      { S7_Templates := "SrcType := Int" } LE_Contact(in1 := "100_GCU_AUTO_SEQ_DB".CRNT_STEP, in2 := 470)
   END_RUNG wire#w1
   // the same network as SCL:
   "Setpoint Override_DB"(Enable := ("100_GCU_AUTO_SEQ_DB".CRNT_STEP >= 290) AND ("100_GCU_AUTO_SEQ_DB".CRNT_STEP <= 470),   // "Setpoint Override"
                          "Activate Temp Prot" := "80_From_HMI"."TT002 Target Protection",
                          Temperature := "12_AI_Data".E_400_TE002_SCALED,
                          "Temperature Setpoint" := "84_Setpoints".E400_TT002_HighHigh,
                          "Temperature Tolerance" := "84_Setpoints"."E-400 TT002 Tolerance",
                          "Activate Press Prot" := "80_From_HMI"."PT002 Target Protection",
                          Pressure := "12_AI_Data".E_400_PT002_SCALED,
                          "Pressure Setpoint" := "84_Setpoints".E400_PT002_High,
                          "Pressure Tolerance" := "84_Setpoints"."E-400 PT002 Tolerance",
                          "Pressure Target" := "84_Setpoints".PIT416_Target,
                          "Pressure Safe Target" := "84_Setpoints".PIT416_Target_Safe,
                          "Activate Tank Change Prot" := "80_From_HMI"."Tank Close Protection",
                          "Tank Change TimeOut" := "84_Setpoints"."Tank Close TimeOut",
                          "Pressure Safe Override" => "84_Setpoints".PIT416_Target_Safe,
                          ENO => #_w1);
   IF #_w1 AND "Setpoint Override_DB"."Set Pressure" THEN
       "19_AUTO_CMNDS_Data".PIT416_CMND_Target := "Setpoint Override_DB"."Pressure Target Override";
   END_IF;
END_REGION

REGION Network 6: PIT416 Target Ramp
   RUNG wire#powerrail
      { S7_Templates := "[SrcType := Real, DestType := DInt]" } Convert(in := "86_Times".PIT416_TRGT_RMP_TIME, out => "68_Sys_Status_Data"."PIT416_TRGT_RMP_TIME D_INT")
      Mul(in1 := "68_Sys_Status_Data"."PIT416_TRGT_RMP_TIME D_INT", in2 := 1000, out => "RAMP_DB"."Time span")
      "RAMP_DB"(Start := wire#w1, "Time span" :=, "Minimum Value" := "12_AI_Data".PIT_416_SCALED, "Maximum Value" := "84_Setpoints".PIT416_Target, Value =>, "Ramp Done" =>)
      I_Contact( "Setpoint Override_DB"."Set Pressure" )
      Move(in := "RAMP_DB".Value, out1 => "19_AUTO_CMNDS_Data".PIT416_CMND_Target)
   END_RUNG
   RUNG wire#powerrail
      { S7_Templates := "SrcType := Int" } GE_Contact(in1 := "100_GCU_AUTO_SEQ_DB".CRNT_STEP, in2 := 290)
      { S7_Templates := "SrcType := Int" } LT_Contact(in1 := "100_GCU_AUTO_SEQ_DB".CRNT_STEP, in2 := 450)
   END_RUNG wire#w1
   // the same network as SCL:
   "68_Sys_Status_Data"."PIT416_TRGT_RMP_TIME D_INT" := REAL_TO_DINT("86_Times".PIT416_TRGT_RMP_TIME);
   "RAMP_DB"."Time span" := "68_Sys_Status_Data"."PIT416_TRGT_RMP_TIME D_INT" * 1000;
   "RAMP_DB"(Start := ("100_GCU_AUTO_SEQ_DB".CRNT_STEP >= 290) AND ("100_GCU_AUTO_SEQ_DB".CRNT_STEP < 450),   // "RAMP"
             "Minimum Value" := "12_AI_Data".PIT_416_SCALED,
             "Maximum Value" := "84_Setpoints".PIT416_Target,
             ENO => #_w1);
   IF #_w1 AND NOT "Setpoint Override_DB"."Set Pressure" THEN
       "19_AUTO_CMNDS_Data".PIT416_CMND_Target := "RAMP_DB".Value;
   END_IF;
END_REGION
END_FUNCTION

FUNCTION "150_GCU_LCL_CNTRL" : Void   // FC150, LAD
TITLE = GCU Local Control
{ S7_Optimized_Access := 'TRUE' }
AUTHOR : JRS
VERSION : 0.1
// For automatic control of the GCU from the HMI and not the BWTS or BTCS
   VAR_TEMP   // added for the SCL form of the ladder/FBD networks
      _w1 : Bool;
   END_VAR
BEGIN

REGION Network 1: System Ok For Local Control
   // Valves at initial etc
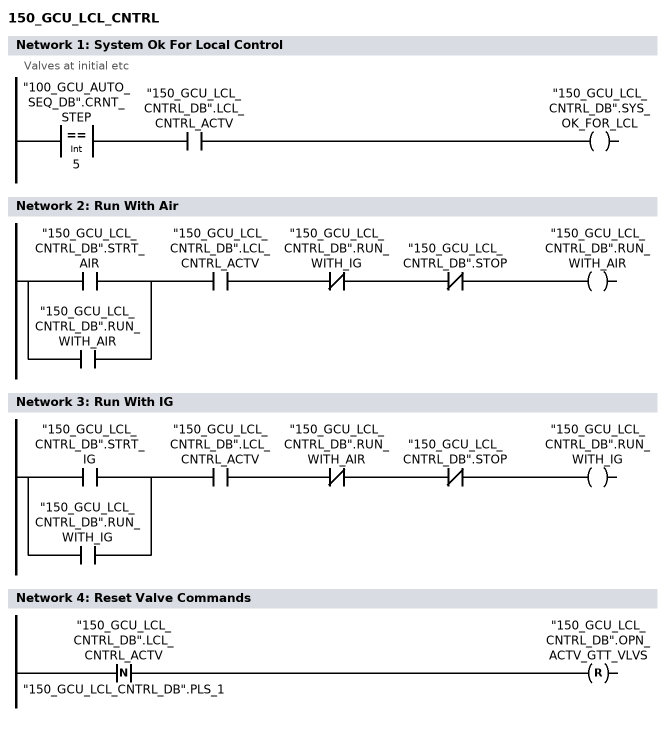
   RUNG wire#powerrail
      { S7_Templates := "SrcType := Int" } EQ_Contact(in1 := "100_GCU_AUTO_SEQ_DB".CRNT_STEP, in2 := 5)
      Contact( "150_GCU_LCL_CNTRL_DB".LCL_CNTRL_ACTV )
      Coil( "150_GCU_LCL_CNTRL_DB".SYS_OK_FOR_LCL )
   END_RUNG
   // the same network as SCL:
   "150_GCU_LCL_CNTRL_DB".SYS_OK_FOR_LCL := ("100_GCU_AUTO_SEQ_DB".CRNT_STEP = 5) AND "150_GCU_LCL_CNTRL_DB".LCL_CNTRL_ACTV;
END_REGION

REGION Network 2: Run With Air
   RUNG wire#powerrail
      Contact( "150_GCU_LCL_CNTRL_DB".STRT_AIR )
      wire#w1
      Contact( "150_GCU_LCL_CNTRL_DB".LCL_CNTRL_ACTV )
      I_Contact( "150_GCU_LCL_CNTRL_DB".RUN_WITH_IG )
      I_Contact( "150_GCU_LCL_CNTRL_DB".STOP )
      Coil( "150_GCU_LCL_CNTRL_DB".RUN_WITH_AIR )
   END_RUNG
   RUNG wire#powerrail
      Contact( "150_GCU_LCL_CNTRL_DB".RUN_WITH_AIR )
   END_RUNG wire#w1
   // the same network as SCL:
   "150_GCU_LCL_CNTRL_DB".RUN_WITH_AIR := ("150_GCU_LCL_CNTRL_DB".STRT_AIR OR "150_GCU_LCL_CNTRL_DB".RUN_WITH_AIR) AND "150_GCU_LCL_CNTRL_DB".LCL_CNTRL_ACTV AND NOT "150_GCU_LCL_CNTRL_DB".RUN_WITH_IG AND NOT "150_GCU_LCL_CNTRL_DB".STOP;
END_REGION

REGION Network 3: Run With IG
   RUNG wire#powerrail
      Contact( "150_GCU_LCL_CNTRL_DB".STRT_IG )
      wire#w1
      Contact( "150_GCU_LCL_CNTRL_DB".LCL_CNTRL_ACTV )
      I_Contact( "150_GCU_LCL_CNTRL_DB".RUN_WITH_AIR )
      I_Contact( "150_GCU_LCL_CNTRL_DB".STOP )
      Coil( "150_GCU_LCL_CNTRL_DB".RUN_WITH_IG )
   END_RUNG
   RUNG wire#powerrail
      Contact( "150_GCU_LCL_CNTRL_DB".RUN_WITH_IG )
   END_RUNG wire#w1
   // the same network as SCL:
   "150_GCU_LCL_CNTRL_DB".RUN_WITH_IG := ("150_GCU_LCL_CNTRL_DB".STRT_IG OR "150_GCU_LCL_CNTRL_DB".RUN_WITH_IG) AND "150_GCU_LCL_CNTRL_DB".LCL_CNTRL_ACTV AND NOT "150_GCU_LCL_CNTRL_DB".RUN_WITH_AIR AND NOT "150_GCU_LCL_CNTRL_DB".STOP;
END_REGION

REGION Network 4: Reset Valve Commands
   RUNG wire#powerrail
      N_Contact(operand := "150_GCU_LCL_CNTRL_DB".LCL_CNTRL_ACTV, bit := "150_GCU_LCL_CNTRL_DB".PLS_1)
      R_Coil( "150_GCU_LCL_CNTRL_DB".OPN_ACTV_GTT_VLVS )
   END_RUNG
   // the same network as SCL:
   #_w1 := NOT "150_GCU_LCL_CNTRL_DB".LCL_CNTRL_ACTV AND "150_GCU_LCL_CNTRL_DB".PLS_1;   // falling edge of "150_GCU_LCL_CNTRL_DB".LCL_CNTRL_ACTV
   "150_GCU_LCL_CNTRL_DB".PLS_1 := "150_GCU_LCL_CNTRL_DB".LCL_CNTRL_ACTV;
   IF #_w1 THEN "150_GCU_LCL_CNTRL_DB".OPN_ACTV_GTT_VLVS := FALSE; END_IF;
END_REGION
END_FUNCTION

// folder: 1000 - 1999 BWT System Control/1060 - 1089 Alarm & Valve Status Handling

FUNCTION "1060_ALARMS_TO_WORDS" : Void   // FC1060, LAD
TITLE = Alarm Processing
{ S7_Optimized_Access := 'TRUE' }
AUTHOR : JRS
VERSION : 0.1
// To determine alarm conditions
BEGIN

REGION Network 1: DB64 DBX18.0 = TX425/426 Tank 1 pH Low Alarm
   // BWTS_ALARM_WORD_10_BIT_0
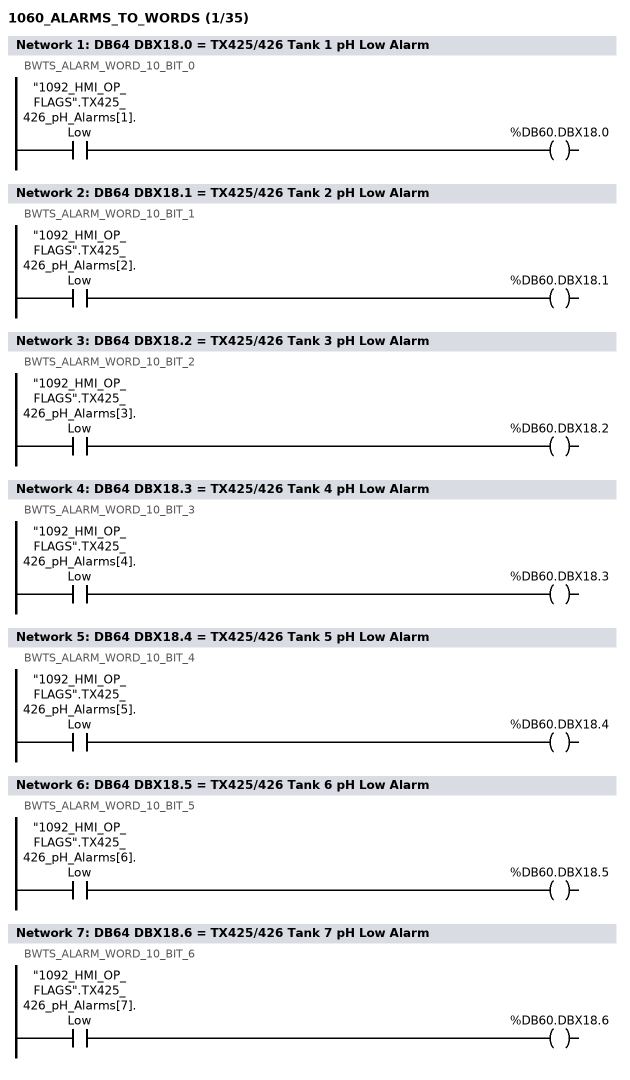
   RUNG wire#powerrail
      Contact( "1092_HMI_OP_FLAGS".TX425_426_pH_Alarms[1].Low )
      Coil( %DB60.DBX18.0 )
   END_RUNG
   // the same network as SCL:
   %DB60.DBX18.0 := "1092_HMI_OP_FLAGS".TX425_426_pH_Alarms[1].Low;
END_REGION

REGION Network 2: DB64 DBX18.1 = TX425/426 Tank 2 pH Low Alarm
   // BWTS_ALARM_WORD_10_BIT_1
   RUNG wire#powerrail
      Contact( "1092_HMI_OP_FLAGS".TX425_426_pH_Alarms[2].Low )
      Coil( %DB60.DBX18.1 )
   END_RUNG
   // the same network as SCL:
   %DB60.DBX18.1 := "1092_HMI_OP_FLAGS".TX425_426_pH_Alarms[2].Low;
END_REGION

REGION Network 3: DB64 DBX18.2 = TX425/426 Tank 3 pH Low Alarm
   // BWTS_ALARM_WORD_10_BIT_2
   RUNG wire#powerrail
      Contact( "1092_HMI_OP_FLAGS".TX425_426_pH_Alarms[3].Low )
      Coil( %DB60.DBX18.2 )
   END_RUNG
   // the same network as SCL:
   %DB60.DBX18.2 := "1092_HMI_OP_FLAGS".TX425_426_pH_Alarms[3].Low;
END_REGION

REGION Network 4: DB64 DBX18.3 = TX425/426 Tank 4 pH Low Alarm
   // BWTS_ALARM_WORD_10_BIT_3
   RUNG wire#powerrail
      Contact( "1092_HMI_OP_FLAGS".TX425_426_pH_Alarms[4].Low )
      Coil( %DB60.DBX18.3 )
   END_RUNG
   // the same network as SCL:
   %DB60.DBX18.3 := "1092_HMI_OP_FLAGS".TX425_426_pH_Alarms[4].Low;
END_REGION

REGION Network 5: DB64 DBX18.4 = TX425/426 Tank 5 pH Low Alarm
   // BWTS_ALARM_WORD_10_BIT_4
   RUNG wire#powerrail
      Contact( "1092_HMI_OP_FLAGS".TX425_426_pH_Alarms[5].Low )
      Coil( %DB60.DBX18.4 )
   END_RUNG
   // the same network as SCL:
   %DB60.DBX18.4 := "1092_HMI_OP_FLAGS".TX425_426_pH_Alarms[5].Low;
END_REGION

REGION Network 6: DB64 DBX18.5 = TX425/426 Tank 6 pH Low Alarm
   // BWTS_ALARM_WORD_10_BIT_5
   RUNG wire#powerrail
      Contact( "1092_HMI_OP_FLAGS".TX425_426_pH_Alarms[6].Low )
      Coil( %DB60.DBX18.5 )
   END_RUNG
   // the same network as SCL:
   %DB60.DBX18.5 := "1092_HMI_OP_FLAGS".TX425_426_pH_Alarms[6].Low;
END_REGION

REGION Network 7: DB64 DBX18.6 = TX425/426 Tank 7 pH Low Alarm
   // BWTS_ALARM_WORD_10_BIT_6
   RUNG wire#powerrail
      Contact( "1092_HMI_OP_FLAGS".TX425_426_pH_Alarms[7].Low )
      Coil( %DB60.DBX18.6 )
   END_RUNG
   // the same network as SCL:
   %DB60.DBX18.6 := "1092_HMI_OP_FLAGS".TX425_426_pH_Alarms[7].Low;
END_REGION

REGION Network 8: DB64 DBX18.7 = TX425/426 Tank 8 pH Low Alarm
   // BWTS_ALARM_WORD_10_BIT_7
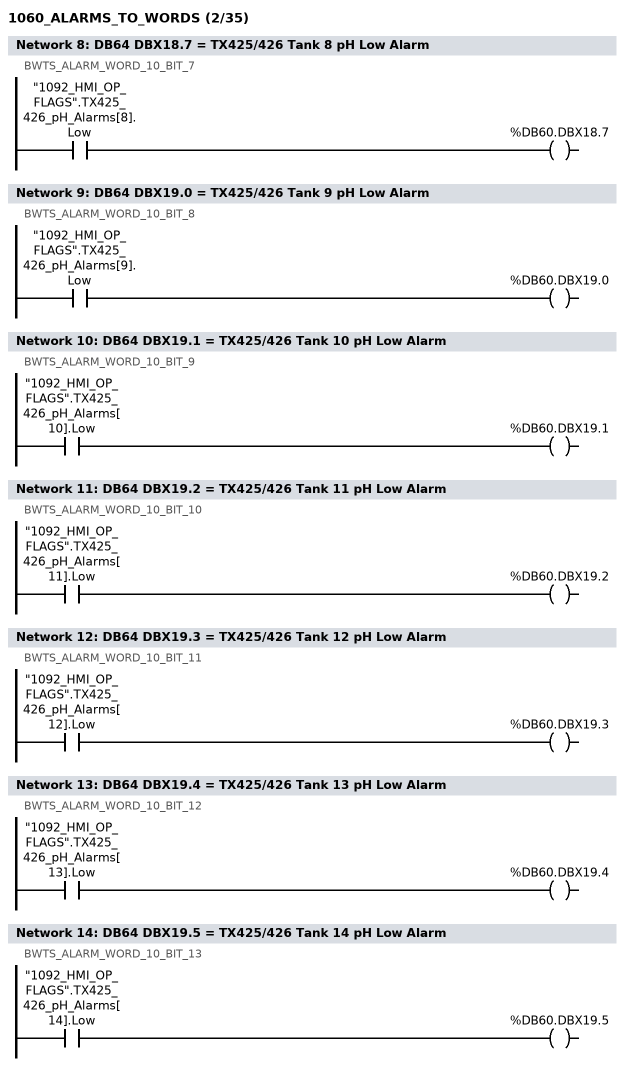
   RUNG wire#powerrail
      Contact( "1092_HMI_OP_FLAGS".TX425_426_pH_Alarms[8].Low )
      Coil( %DB60.DBX18.7 )
   END_RUNG
   // the same network as SCL:
   %DB60.DBX18.7 := "1092_HMI_OP_FLAGS".TX425_426_pH_Alarms[8].Low;
END_REGION

REGION Network 9: DB64 DBX19.0 = TX425/426 Tank 9 pH Low Alarm
   // BWTS_ALARM_WORD_10_BIT_8
   RUNG wire#powerrail
      Contact( "1092_HMI_OP_FLAGS".TX425_426_pH_Alarms[9].Low )
      Coil( %DB60.DBX19.0 )
   END_RUNG
   // the same network as SCL:
   %DB60.DBX19.0 := "1092_HMI_OP_FLAGS".TX425_426_pH_Alarms[9].Low;
END_REGION

REGION Network 10: DB64 DBX19.1 = TX425/426 Tank 10 pH Low Alarm
   // BWTS_ALARM_WORD_10_BIT_9
   RUNG wire#powerrail
      Contact( "1092_HMI_OP_FLAGS".TX425_426_pH_Alarms[10].Low )
      Coil( %DB60.DBX19.1 )
   END_RUNG
   // the same network as SCL:
   %DB60.DBX19.1 := "1092_HMI_OP_FLAGS".TX425_426_pH_Alarms[10].Low;
END_REGION

REGION Network 11: DB64 DBX19.2 = TX425/426 Tank 11 pH Low Alarm
   // BWTS_ALARM_WORD_10_BIT_10
   RUNG wire#powerrail
      Contact( "1092_HMI_OP_FLAGS".TX425_426_pH_Alarms[11].Low )
      Coil( %DB60.DBX19.2 )
   END_RUNG
   // the same network as SCL:
   %DB60.DBX19.2 := "1092_HMI_OP_FLAGS".TX425_426_pH_Alarms[11].Low;
END_REGION

REGION Network 12: DB64 DBX19.3 = TX425/426 Tank 12 pH Low Alarm
   // BWTS_ALARM_WORD_10_BIT_11
   RUNG wire#powerrail
      Contact( "1092_HMI_OP_FLAGS".TX425_426_pH_Alarms[12].Low )
      Coil( %DB60.DBX19.3 )
   END_RUNG
   // the same network as SCL:
   %DB60.DBX19.3 := "1092_HMI_OP_FLAGS".TX425_426_pH_Alarms[12].Low;
END_REGION

REGION Network 13: DB64 DBX19.4 = TX425/426 Tank 13 pH Low Alarm
   // BWTS_ALARM_WORD_10_BIT_12
   RUNG wire#powerrail
      Contact( "1092_HMI_OP_FLAGS".TX425_426_pH_Alarms[13].Low )
      Coil( %DB60.DBX19.4 )
   END_RUNG
   // the same network as SCL:
   %DB60.DBX19.4 := "1092_HMI_OP_FLAGS".TX425_426_pH_Alarms[13].Low;
END_REGION

REGION Network 14: DB64 DBX19.5 = TX425/426 Tank 14 pH Low Alarm
   // BWTS_ALARM_WORD_10_BIT_13
   RUNG wire#powerrail
      Contact( "1092_HMI_OP_FLAGS".TX425_426_pH_Alarms[14].Low )
      Coil( %DB60.DBX19.5 )
   END_RUNG
   // the same network as SCL:
   %DB60.DBX19.5 := "1092_HMI_OP_FLAGS".TX425_426_pH_Alarms[14].Low;
END_REGION

REGION Network 16: DB64 DBX20.0 = TX427/428 Tank 1 DO Low Alarm
   // BWTS_ALARM_WORD_11_BIT_0
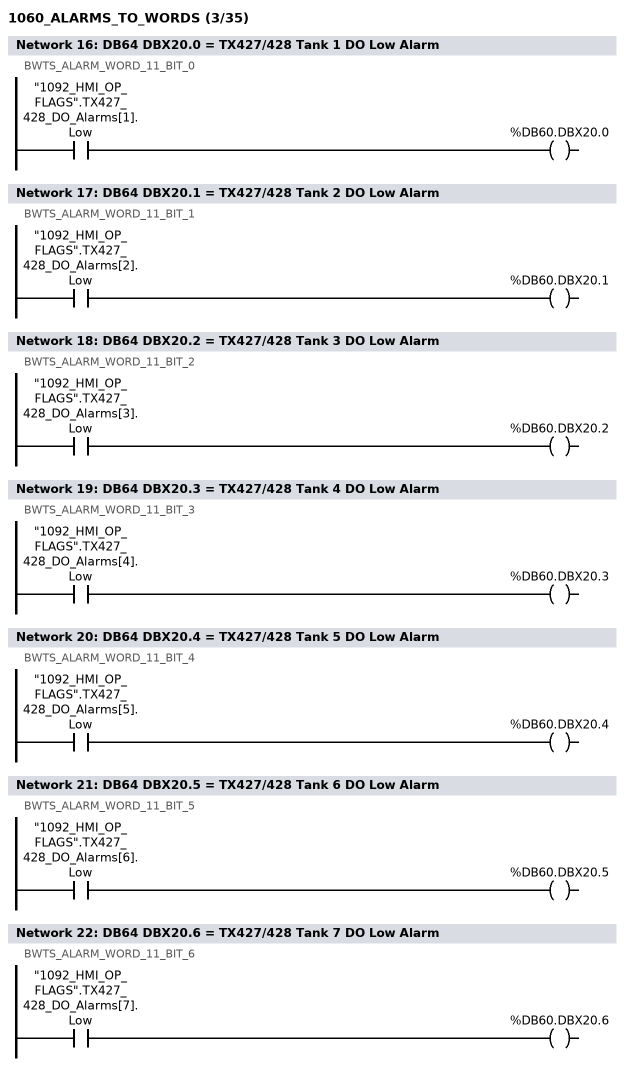
   RUNG wire#powerrail
      Contact( "1092_HMI_OP_FLAGS".TX427_428_DO_Alarms[1].Low )
      Coil( %DB60.DBX20.0 )
   END_RUNG
   // the same network as SCL:
   %DB60.DBX20.0 := "1092_HMI_OP_FLAGS".TX427_428_DO_Alarms[1].Low;
END_REGION

REGION Network 17: DB64 DBX20.1 = TX427/428 Tank 2 DO Low Alarm
   // BWTS_ALARM_WORD_11_BIT_1
   RUNG wire#powerrail
      Contact( "1092_HMI_OP_FLAGS".TX427_428_DO_Alarms[2].Low )
      Coil( %DB60.DBX20.1 )
   END_RUNG
   // the same network as SCL:
   %DB60.DBX20.1 := "1092_HMI_OP_FLAGS".TX427_428_DO_Alarms[2].Low;
END_REGION

REGION Network 18: DB64 DBX20.2 = TX427/428 Tank 3 DO Low Alarm
   // BWTS_ALARM_WORD_11_BIT_2
   RUNG wire#powerrail
      Contact( "1092_HMI_OP_FLAGS".TX427_428_DO_Alarms[3].Low )
      Coil( %DB60.DBX20.2 )
   END_RUNG
   // the same network as SCL:
   %DB60.DBX20.2 := "1092_HMI_OP_FLAGS".TX427_428_DO_Alarms[3].Low;
END_REGION

REGION Network 19: DB64 DBX20.3 = TX427/428 Tank 4 DO Low Alarm
   // BWTS_ALARM_WORD_11_BIT_3
   RUNG wire#powerrail
      Contact( "1092_HMI_OP_FLAGS".TX427_428_DO_Alarms[4].Low )
      Coil( %DB60.DBX20.3 )
   END_RUNG
   // the same network as SCL:
   %DB60.DBX20.3 := "1092_HMI_OP_FLAGS".TX427_428_DO_Alarms[4].Low;
END_REGION

REGION Network 20: DB64 DBX20.4 = TX427/428 Tank 5 DO Low Alarm
   // BWTS_ALARM_WORD_11_BIT_4
   RUNG wire#powerrail
      Contact( "1092_HMI_OP_FLAGS".TX427_428_DO_Alarms[5].Low )
      Coil( %DB60.DBX20.4 )
   END_RUNG
   // the same network as SCL:
   %DB60.DBX20.4 := "1092_HMI_OP_FLAGS".TX427_428_DO_Alarms[5].Low;
END_REGION

REGION Network 21: DB64 DBX20.5 = TX427/428 Tank 6 DO Low Alarm
   // BWTS_ALARM_WORD_11_BIT_5
   RUNG wire#powerrail
      Contact( "1092_HMI_OP_FLAGS".TX427_428_DO_Alarms[6].Low )
      Coil( %DB60.DBX20.5 )
   END_RUNG
   // the same network as SCL:
   %DB60.DBX20.5 := "1092_HMI_OP_FLAGS".TX427_428_DO_Alarms[6].Low;
END_REGION

REGION Network 22: DB64 DBX20.6 = TX427/428 Tank 7 DO Low Alarm
   // BWTS_ALARM_WORD_11_BIT_6
   RUNG wire#powerrail
      Contact( "1092_HMI_OP_FLAGS".TX427_428_DO_Alarms[7].Low )
      Coil( %DB60.DBX20.6 )
   END_RUNG
   // the same network as SCL:
   %DB60.DBX20.6 := "1092_HMI_OP_FLAGS".TX427_428_DO_Alarms[7].Low;
END_REGION

REGION Network 23: DB64 DBX20.7 = TX427/428 Tank 8 DO Low Alarm
   // BWTS_ALARM_WORD_11_BIT_7
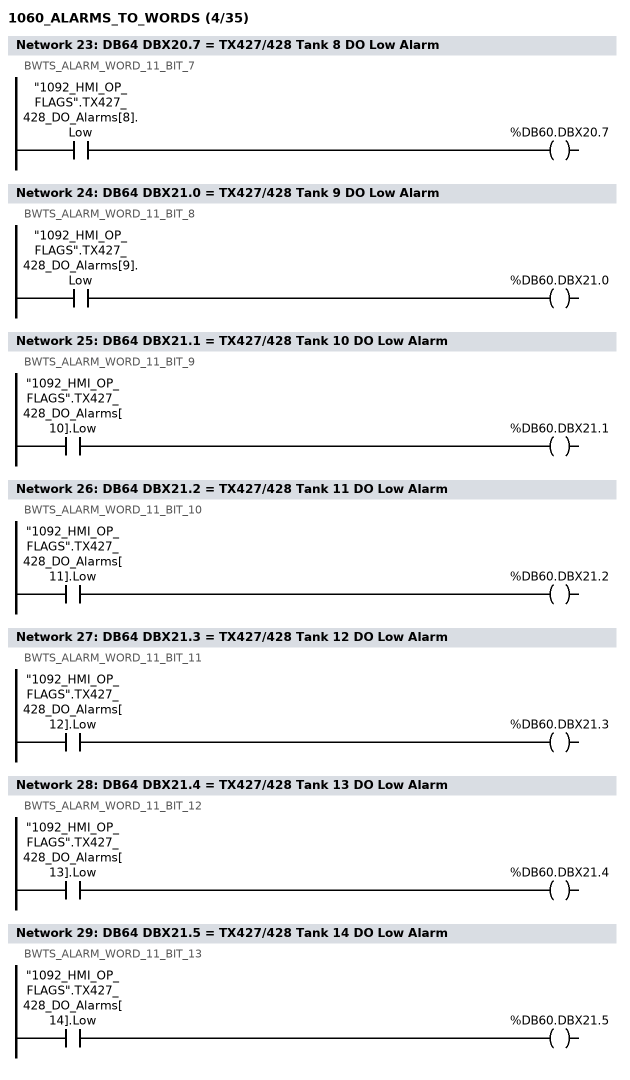
   RUNG wire#powerrail
      Contact( "1092_HMI_OP_FLAGS".TX427_428_DO_Alarms[8].Low )
      Coil( %DB60.DBX20.7 )
   END_RUNG
   // the same network as SCL:
   %DB60.DBX20.7 := "1092_HMI_OP_FLAGS".TX427_428_DO_Alarms[8].Low;
END_REGION

REGION Network 24: DB64 DBX21.0 = TX427/428 Tank 9 DO Low Alarm
   // BWTS_ALARM_WORD_11_BIT_8
   RUNG wire#powerrail
      Contact( "1092_HMI_OP_FLAGS".TX427_428_DO_Alarms[9].Low )
      Coil( %DB60.DBX21.0 )
   END_RUNG
   // the same network as SCL:
   %DB60.DBX21.0 := "1092_HMI_OP_FLAGS".TX427_428_DO_Alarms[9].Low;
END_REGION

REGION Network 25: DB64 DBX21.1 = TX427/428 Tank 10 DO Low Alarm
   // BWTS_ALARM_WORD_11_BIT_9
   RUNG wire#powerrail
      Contact( "1092_HMI_OP_FLAGS".TX427_428_DO_Alarms[10].Low )
      Coil( %DB60.DBX21.1 )
   END_RUNG
   // the same network as SCL:
   %DB60.DBX21.1 := "1092_HMI_OP_FLAGS".TX427_428_DO_Alarms[10].Low;
END_REGION

REGION Network 26: DB64 DBX21.2 = TX427/428 Tank 11 DO Low Alarm
   // BWTS_ALARM_WORD_11_BIT_10
   RUNG wire#powerrail
      Contact( "1092_HMI_OP_FLAGS".TX427_428_DO_Alarms[11].Low )
      Coil( %DB60.DBX21.2 )
   END_RUNG
   // the same network as SCL:
   %DB60.DBX21.2 := "1092_HMI_OP_FLAGS".TX427_428_DO_Alarms[11].Low;
END_REGION

REGION Network 27: DB64 DBX21.3 = TX427/428 Tank 12 DO Low Alarm
   // BWTS_ALARM_WORD_11_BIT_11
   RUNG wire#powerrail
      Contact( "1092_HMI_OP_FLAGS".TX427_428_DO_Alarms[12].Low )
      Coil( %DB60.DBX21.3 )
   END_RUNG
   // the same network as SCL:
   %DB60.DBX21.3 := "1092_HMI_OP_FLAGS".TX427_428_DO_Alarms[12].Low;
END_REGION

REGION Network 28: DB64 DBX21.4 = TX427/428 Tank 13 DO Low Alarm
   // BWTS_ALARM_WORD_11_BIT_12
   RUNG wire#powerrail
      Contact( "1092_HMI_OP_FLAGS".TX427_428_DO_Alarms[13].Low )
      Coil( %DB60.DBX21.4 )
   END_RUNG
   // the same network as SCL:
   %DB60.DBX21.4 := "1092_HMI_OP_FLAGS".TX427_428_DO_Alarms[13].Low;
END_REGION

REGION Network 29: DB64 DBX21.5 = TX427/428 Tank 14 DO Low Alarm
   // BWTS_ALARM_WORD_11_BIT_13
   RUNG wire#powerrail
      Contact( "1092_HMI_OP_FLAGS".TX427_428_DO_Alarms[14].Low )
      Coil( %DB60.DBX21.5 )
   END_RUNG
   // the same network as SCL:
   %DB60.DBX21.5 := "1092_HMI_OP_FLAGS".TX427_428_DO_Alarms[14].Low;
END_REGION

REGION Network 31: DB64 DBX22.0 = USD Flow Tank 1 Low Low
   // BWTS_ALARM_WORD_12_BIT_0
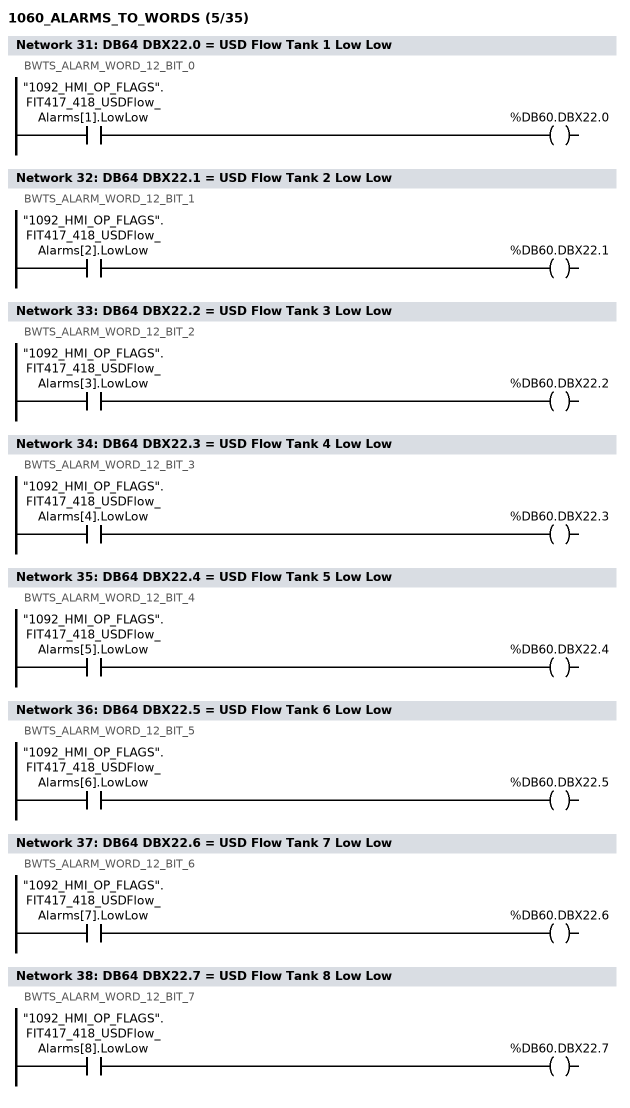
   RUNG wire#powerrail
      Contact( "1092_HMI_OP_FLAGS".FIT417_418_USDFlow_Alarms[1].LowLow )
      Coil( %DB60.DBX22.0 )
   END_RUNG
   // the same network as SCL:
   %DB60.DBX22.0 := "1092_HMI_OP_FLAGS".FIT417_418_USDFlow_Alarms[1].LowLow;
END_REGION

REGION Network 32: DB64 DBX22.1 = USD Flow Tank 2 Low Low
   // BWTS_ALARM_WORD_12_BIT_1
   RUNG wire#powerrail
      Contact( "1092_HMI_OP_FLAGS".FIT417_418_USDFlow_Alarms[2].LowLow )
      Coil( %DB60.DBX22.1 )
   END_RUNG
   // the same network as SCL:
   %DB60.DBX22.1 := "1092_HMI_OP_FLAGS".FIT417_418_USDFlow_Alarms[2].LowLow;
END_REGION

REGION Network 33: DB64 DBX22.2 = USD Flow Tank 3 Low Low
   // BWTS_ALARM_WORD_12_BIT_2
   RUNG wire#powerrail
      Contact( "1092_HMI_OP_FLAGS".FIT417_418_USDFlow_Alarms[3].LowLow )
      Coil( %DB60.DBX22.2 )
   END_RUNG
   // the same network as SCL:
   %DB60.DBX22.2 := "1092_HMI_OP_FLAGS".FIT417_418_USDFlow_Alarms[3].LowLow;
END_REGION

REGION Network 34: DB64 DBX22.3 = USD Flow Tank 4 Low Low
   // BWTS_ALARM_WORD_12_BIT_3
   RUNG wire#powerrail
      Contact( "1092_HMI_OP_FLAGS".FIT417_418_USDFlow_Alarms[4].LowLow )
      Coil( %DB60.DBX22.3 )
   END_RUNG
   // the same network as SCL:
   %DB60.DBX22.3 := "1092_HMI_OP_FLAGS".FIT417_418_USDFlow_Alarms[4].LowLow;
END_REGION

REGION Network 35: DB64 DBX22.4 = USD Flow Tank 5 Low Low
   // BWTS_ALARM_WORD_12_BIT_4
   RUNG wire#powerrail
      Contact( "1092_HMI_OP_FLAGS".FIT417_418_USDFlow_Alarms[5].LowLow )
      Coil( %DB60.DBX22.4 )
   END_RUNG
   // the same network as SCL:
   %DB60.DBX22.4 := "1092_HMI_OP_FLAGS".FIT417_418_USDFlow_Alarms[5].LowLow;
END_REGION

REGION Network 36: DB64 DBX22.5 = USD Flow Tank 6 Low Low
   // BWTS_ALARM_WORD_12_BIT_5
   RUNG wire#powerrail
      Contact( "1092_HMI_OP_FLAGS".FIT417_418_USDFlow_Alarms[6].LowLow )
      Coil( %DB60.DBX22.5 )
   END_RUNG
   // the same network as SCL:
   %DB60.DBX22.5 := "1092_HMI_OP_FLAGS".FIT417_418_USDFlow_Alarms[6].LowLow;
END_REGION

REGION Network 37: DB64 DBX22.6 = USD Flow Tank 7 Low Low
   // BWTS_ALARM_WORD_12_BIT_6
   RUNG wire#powerrail
      Contact( "1092_HMI_OP_FLAGS".FIT417_418_USDFlow_Alarms[7].LowLow )
      Coil( %DB60.DBX22.6 )
   END_RUNG
   // the same network as SCL:
   %DB60.DBX22.6 := "1092_HMI_OP_FLAGS".FIT417_418_USDFlow_Alarms[7].LowLow;
END_REGION

REGION Network 38: DB64 DBX22.7 = USD Flow Tank 8 Low Low
   // BWTS_ALARM_WORD_12_BIT_7
   RUNG wire#powerrail
      Contact( "1092_HMI_OP_FLAGS".FIT417_418_USDFlow_Alarms[8].LowLow )
      Coil( %DB60.DBX22.7 )
   END_RUNG
   // the same network as SCL:
   %DB60.DBX22.7 := "1092_HMI_OP_FLAGS".FIT417_418_USDFlow_Alarms[8].LowLow;
END_REGION

REGION Network 39: DB64 DBX23.0 = USD Flow Tank 9 Low Low
   // BWTS_ALARM_WORD_12_BIT_8
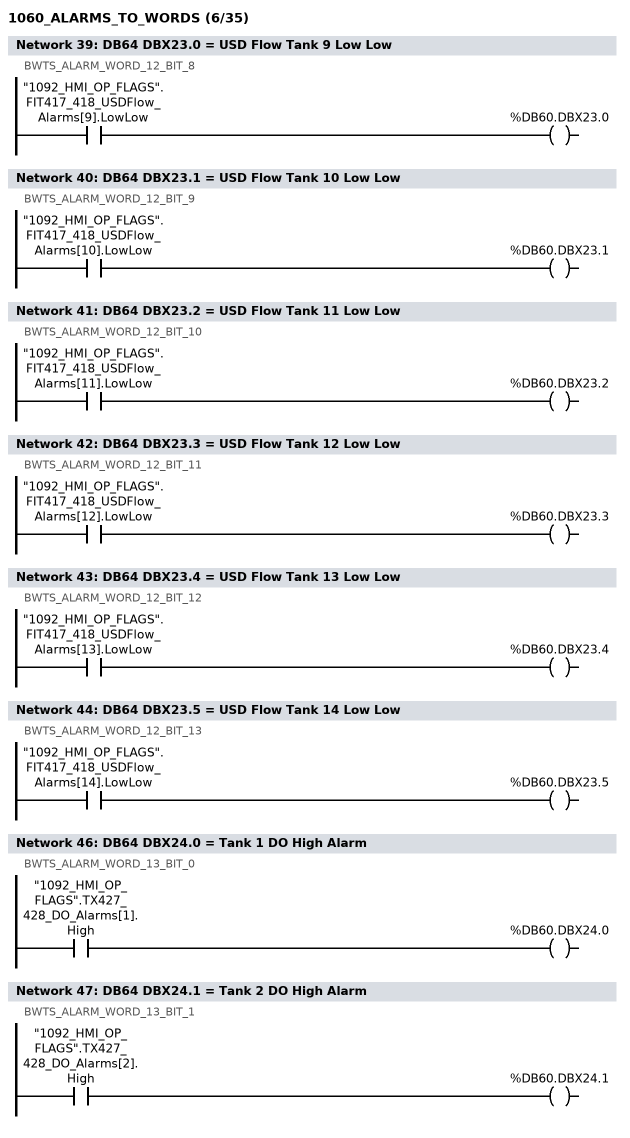
   RUNG wire#powerrail
      Contact( "1092_HMI_OP_FLAGS".FIT417_418_USDFlow_Alarms[9].LowLow )
      Coil( %DB60.DBX23.0 )
   END_RUNG
   // the same network as SCL:
   %DB60.DBX23.0 := "1092_HMI_OP_FLAGS".FIT417_418_USDFlow_Alarms[9].LowLow;
END_REGION

REGION Network 40: DB64 DBX23.1 = USD Flow Tank 10 Low Low
   // BWTS_ALARM_WORD_12_BIT_9
   RUNG wire#powerrail
      Contact( "1092_HMI_OP_FLAGS".FIT417_418_USDFlow_Alarms[10].LowLow )
      Coil( %DB60.DBX23.1 )
   END_RUNG
   // the same network as SCL:
   %DB60.DBX23.1 := "1092_HMI_OP_FLAGS".FIT417_418_USDFlow_Alarms[10].LowLow;
END_REGION

REGION Network 41: DB64 DBX23.2 = USD Flow Tank 11 Low Low
   // BWTS_ALARM_WORD_12_BIT_10
   RUNG wire#powerrail
      Contact( "1092_HMI_OP_FLAGS".FIT417_418_USDFlow_Alarms[11].LowLow )
      Coil( %DB60.DBX23.2 )
   END_RUNG
   // the same network as SCL:
   %DB60.DBX23.2 := "1092_HMI_OP_FLAGS".FIT417_418_USDFlow_Alarms[11].LowLow;
END_REGION

REGION Network 42: DB64 DBX23.3 = USD Flow Tank 12 Low Low
   // BWTS_ALARM_WORD_12_BIT_11
   RUNG wire#powerrail
      Contact( "1092_HMI_OP_FLAGS".FIT417_418_USDFlow_Alarms[12].LowLow )
      Coil( %DB60.DBX23.3 )
   END_RUNG
   // the same network as SCL:
   %DB60.DBX23.3 := "1092_HMI_OP_FLAGS".FIT417_418_USDFlow_Alarms[12].LowLow;
END_REGION

REGION Network 43: DB64 DBX23.4 = USD Flow Tank 13 Low Low
   // BWTS_ALARM_WORD_12_BIT_12
   RUNG wire#powerrail
      Contact( "1092_HMI_OP_FLAGS".FIT417_418_USDFlow_Alarms[13].LowLow )
      Coil( %DB60.DBX23.4 )
   END_RUNG
   // the same network as SCL:
   %DB60.DBX23.4 := "1092_HMI_OP_FLAGS".FIT417_418_USDFlow_Alarms[13].LowLow;
END_REGION

REGION Network 44: DB64 DBX23.5 = USD Flow Tank 14 Low Low
   // BWTS_ALARM_WORD_12_BIT_13
   RUNG wire#powerrail
      Contact( "1092_HMI_OP_FLAGS".FIT417_418_USDFlow_Alarms[14].LowLow )
      Coil( %DB60.DBX23.5 )
   END_RUNG
   // the same network as SCL:
   %DB60.DBX23.5 := "1092_HMI_OP_FLAGS".FIT417_418_USDFlow_Alarms[14].LowLow;
END_REGION

REGION Network 46: DB64 DBX24.0 = Tank 1 DO High Alarm
   // BWTS_ALARM_WORD_13_BIT_0
   RUNG wire#powerrail
      Contact( "1092_HMI_OP_FLAGS".TX427_428_DO_Alarms[1].High )
      Coil( %DB60.DBX24.0 )
   END_RUNG
   // the same network as SCL:
   %DB60.DBX24.0 := "1092_HMI_OP_FLAGS".TX427_428_DO_Alarms[1].High;
END_REGION

REGION Network 47: DB64 DBX24.1 = Tank 2 DO High Alarm
   // BWTS_ALARM_WORD_13_BIT_1
   RUNG wire#powerrail
      Contact( "1092_HMI_OP_FLAGS".TX427_428_DO_Alarms[2].High )
      Coil( %DB60.DBX24.1 )
   END_RUNG
   // the same network as SCL:
   %DB60.DBX24.1 := "1092_HMI_OP_FLAGS".TX427_428_DO_Alarms[2].High;
END_REGION

REGION Network 48: DB64 DBX24.2 = Tank 3 DO High Alarm
   // BWTS_ALARM_WORD_13_BIT_2
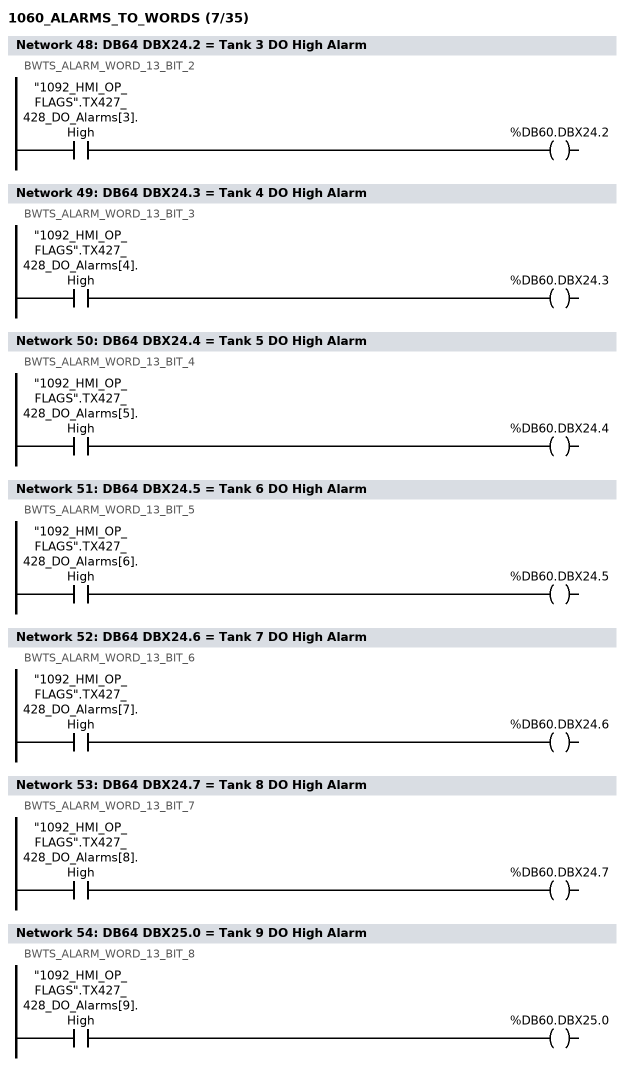
   RUNG wire#powerrail
      Contact( "1092_HMI_OP_FLAGS".TX427_428_DO_Alarms[3].High )
      Coil( %DB60.DBX24.2 )
   END_RUNG
   // the same network as SCL:
   %DB60.DBX24.2 := "1092_HMI_OP_FLAGS".TX427_428_DO_Alarms[3].High;
END_REGION

REGION Network 49: DB64 DBX24.3 = Tank 4 DO High Alarm
   // BWTS_ALARM_WORD_13_BIT_3
   RUNG wire#powerrail
      Contact( "1092_HMI_OP_FLAGS".TX427_428_DO_Alarms[4].High )
      Coil( %DB60.DBX24.3 )
   END_RUNG
   // the same network as SCL:
   %DB60.DBX24.3 := "1092_HMI_OP_FLAGS".TX427_428_DO_Alarms[4].High;
END_REGION

REGION Network 50: DB64 DBX24.4 = Tank 5 DO High Alarm
   // BWTS_ALARM_WORD_13_BIT_4
   RUNG wire#powerrail
      Contact( "1092_HMI_OP_FLAGS".TX427_428_DO_Alarms[5].High )
      Coil( %DB60.DBX24.4 )
   END_RUNG
   // the same network as SCL:
   %DB60.DBX24.4 := "1092_HMI_OP_FLAGS".TX427_428_DO_Alarms[5].High;
END_REGION

REGION Network 51: DB64 DBX24.5 = Tank 6 DO High Alarm
   // BWTS_ALARM_WORD_13_BIT_5
   RUNG wire#powerrail
      Contact( "1092_HMI_OP_FLAGS".TX427_428_DO_Alarms[6].High )
      Coil( %DB60.DBX24.5 )
   END_RUNG
   // the same network as SCL:
   %DB60.DBX24.5 := "1092_HMI_OP_FLAGS".TX427_428_DO_Alarms[6].High;
END_REGION

REGION Network 52: DB64 DBX24.6 = Tank 7 DO High Alarm
   // BWTS_ALARM_WORD_13_BIT_6
   RUNG wire#powerrail
      Contact( "1092_HMI_OP_FLAGS".TX427_428_DO_Alarms[7].High )
      Coil( %DB60.DBX24.6 )
   END_RUNG
   // the same network as SCL:
   %DB60.DBX24.6 := "1092_HMI_OP_FLAGS".TX427_428_DO_Alarms[7].High;
END_REGION

REGION Network 53: DB64 DBX24.7 = Tank 8 DO High Alarm
   // BWTS_ALARM_WORD_13_BIT_7
   RUNG wire#powerrail
      Contact( "1092_HMI_OP_FLAGS".TX427_428_DO_Alarms[8].High )
      Coil( %DB60.DBX24.7 )
   END_RUNG
   // the same network as SCL:
   %DB60.DBX24.7 := "1092_HMI_OP_FLAGS".TX427_428_DO_Alarms[8].High;
END_REGION

REGION Network 54: DB64 DBX25.0 = Tank 9 DO High Alarm
   // BWTS_ALARM_WORD_13_BIT_8
   RUNG wire#powerrail
      Contact( "1092_HMI_OP_FLAGS".TX427_428_DO_Alarms[9].High )
      Coil( %DB60.DBX25.0 )
   END_RUNG
   // the same network as SCL:
   %DB60.DBX25.0 := "1092_HMI_OP_FLAGS".TX427_428_DO_Alarms[9].High;
END_REGION

REGION Network 55: DB64 DBX25.1 = Tank 10 DO High Alarm
   // BWTS_ALARM_WORD_13_BIT_9
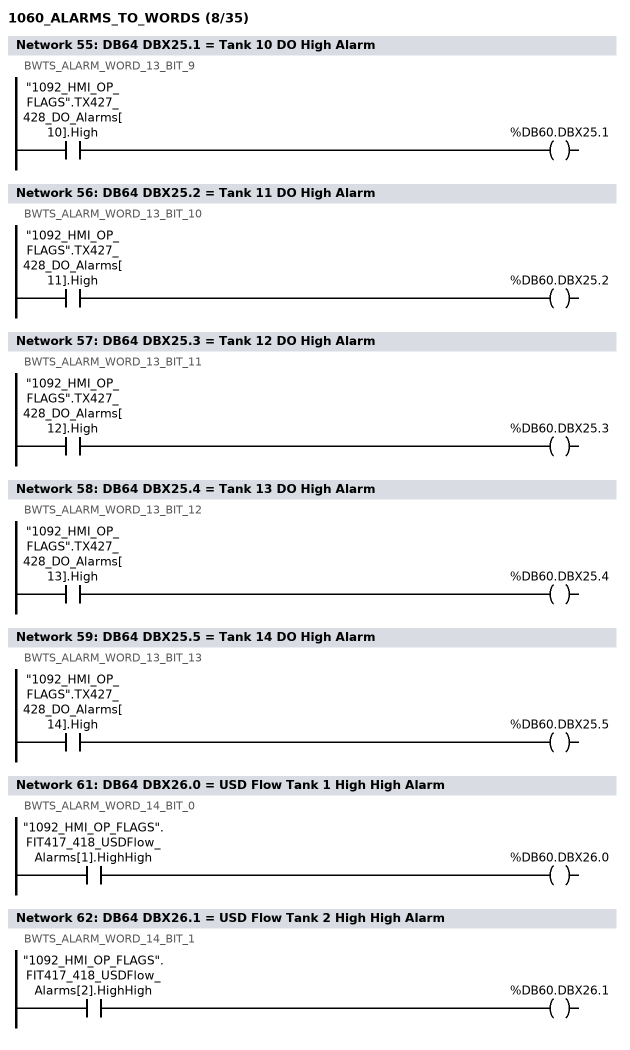
   RUNG wire#powerrail
      Contact( "1092_HMI_OP_FLAGS".TX427_428_DO_Alarms[10].High )
      Coil( %DB60.DBX25.1 )
   END_RUNG
   // the same network as SCL:
   %DB60.DBX25.1 := "1092_HMI_OP_FLAGS".TX427_428_DO_Alarms[10].High;
END_REGION

REGION Network 56: DB64 DBX25.2 = Tank 11 DO High Alarm
   // BWTS_ALARM_WORD_13_BIT_10
   RUNG wire#powerrail
      Contact( "1092_HMI_OP_FLAGS".TX427_428_DO_Alarms[11].High )
      Coil( %DB60.DBX25.2 )
   END_RUNG
   // the same network as SCL:
   %DB60.DBX25.2 := "1092_HMI_OP_FLAGS".TX427_428_DO_Alarms[11].High;
END_REGION

REGION Network 57: DB64 DBX25.3 = Tank 12 DO High Alarm
   // BWTS_ALARM_WORD_13_BIT_11
   RUNG wire#powerrail
      Contact( "1092_HMI_OP_FLAGS".TX427_428_DO_Alarms[12].High )
      Coil( %DB60.DBX25.3 )
   END_RUNG
   // the same network as SCL:
   %DB60.DBX25.3 := "1092_HMI_OP_FLAGS".TX427_428_DO_Alarms[12].High;
END_REGION

REGION Network 58: DB64 DBX25.4 = Tank 13 DO High Alarm
   // BWTS_ALARM_WORD_13_BIT_12
   RUNG wire#powerrail
      Contact( "1092_HMI_OP_FLAGS".TX427_428_DO_Alarms[13].High )
      Coil( %DB60.DBX25.4 )
   END_RUNG
   // the same network as SCL:
   %DB60.DBX25.4 := "1092_HMI_OP_FLAGS".TX427_428_DO_Alarms[13].High;
END_REGION

REGION Network 59: DB64 DBX25.5 = Tank 14 DO High Alarm
   // BWTS_ALARM_WORD_13_BIT_13
   RUNG wire#powerrail
      Contact( "1092_HMI_OP_FLAGS".TX427_428_DO_Alarms[14].High )
      Coil( %DB60.DBX25.5 )
   END_RUNG
   // the same network as SCL:
   %DB60.DBX25.5 := "1092_HMI_OP_FLAGS".TX427_428_DO_Alarms[14].High;
END_REGION

REGION Network 61: DB64 DBX26.0 = USD Flow Tank 1 High High Alarm
   // BWTS_ALARM_WORD_14_BIT_0
   RUNG wire#powerrail
      Contact( "1092_HMI_OP_FLAGS".FIT417_418_USDFlow_Alarms[1].HighHigh )
      Coil( %DB60.DBX26.0 )
   END_RUNG
   // the same network as SCL:
   %DB60.DBX26.0 := "1092_HMI_OP_FLAGS".FIT417_418_USDFlow_Alarms[1].HighHigh;
END_REGION

REGION Network 62: DB64 DBX26.1 = USD Flow Tank 2 High High Alarm
   // BWTS_ALARM_WORD_14_BIT_1
   RUNG wire#powerrail
      Contact( "1092_HMI_OP_FLAGS".FIT417_418_USDFlow_Alarms[2].HighHigh )
      Coil( %DB60.DBX26.1 )
   END_RUNG
   // the same network as SCL:
   %DB60.DBX26.1 := "1092_HMI_OP_FLAGS".FIT417_418_USDFlow_Alarms[2].HighHigh;
END_REGION

REGION Network 63: DB64 DBX26.2 = USD Flow Tank 3 High High Alarm
   // BWTS_ALARM_WORD_14_BIT_2